REGION Network 2
   RUNG wire#powerrail
      { S7_GenerateENO := "TRUE" } Move(in := "1#煤粉仓2#温度":P, out1 => "MNL"."1#煤粉仓2#温度")
   END_RUNG
   // the same network as SCL:
   "MNL"."1#煤粉仓2#温度" := "1#煤粉仓2#温度":P;
END_REGION

REGION Network 3
   RUNG wire#powerrail
      { S7_GenerateENO := "TRUE" } Move(in := "1#煤粉仓3#温度":P, out1 => "MNL"."1#煤粉仓3#温度")
   END_RUNG
   // the same network as SCL:
   "MNL"."1#煤粉仓3#温度" := "1#煤粉仓3#温度":P;
END_REGION

REGION Network 4
   RUNG wire#powerrail
      { S7_GenerateENO := "TRUE" } Move(in := "Tag_101":P, out1 => "MNL"."1#煤粉仓4#温度")
   END_RUNG
   // the same network as SCL:
   "MNL"."1#煤粉仓4#温度" := "Tag_101":P;
END_REGION

REGION Network 5
   RUNG wire#powerrail
      { S7_GenerateENO := "TRUE" } Move(in := "1#煤粉仓5#温度":P, out1 => "MNL"."1#煤粉仓5#温度")
   END_RUNG
   // the same network as SCL:
   "MNL"."1#煤粉仓5#温度" := "1#煤粉仓5#温度":P;
END_REGION

REGION Network 6
   RUNG wire#powerrail
      { S7_GenerateENO := "TRUE" } Move(in := "1#煤粉仓6#温度":P, out1 => "MNL"."1#煤粉仓6#温度")
   END_RUNG
   // the same network as SCL:
   "MNL"."1#煤粉仓6#温度" := "1#煤粉仓6#温度":P;
END_REGION

REGION Network 7
   RUNG wire#powerrail
      { S7_GenerateENO := "TRUE" } Move(in := "2#煤粉仓1#温度":P, out1 => "MNL"."2#煤粉仓1#温度")
   END_RUNG
   // the same network as SCL:
   "MNL"."2#煤粉仓1#温度" := "2#煤粉仓1#温度":P;
END_REGION

REGION Network 8
   RUNG wire#powerrail
      { S7_GenerateENO := "TRUE" } Move(in := "2#煤粉仓2#温度":P, out1 => "MNL"."2#煤粉仓2#温度")
   END_RUNG
   // the same network as SCL:
   "MNL"."2#煤粉仓2#温度" := "2#煤粉仓2#温度":P;
END_REGION

REGION Network 9
   RUNG wire#powerrail
      { S7_GenerateENO := "TRUE" } Move(in := "2#煤粉仓3#温度":P, out1 => "MNL"."2#煤粉仓3#温度")
   END_RUNG
   // the same network as SCL:
   "MNL"."2#煤粉仓3#温度" := "2#煤粉仓3#温度":P;
END_REGION

REGION Network 10
   RUNG wire#powerrail
      { S7_GenerateENO := "TRUE" } Move(in := "2#煤粉仓4#温度":P, out1 => "MNL"."2#煤粉仓4#温度")
   END_RUNG
   // the same network as SCL:
   "MNL"."2#煤粉仓4#温度" := "2#煤粉仓4#温度":P;
END_REGION

REGION Network 11
   RUNG wire#powerrail
      { S7_GenerateENO := "TRUE" } Move(in := "2#煤粉仓5#温度":P, out1 => "MNL"."2#煤粉仓5#温度")
   END_RUNG
   // the same network as SCL:
   "MNL"."2#煤粉仓5#温度" := "2#煤粉仓5#温度":P;
END_REGION

REGION Network 12
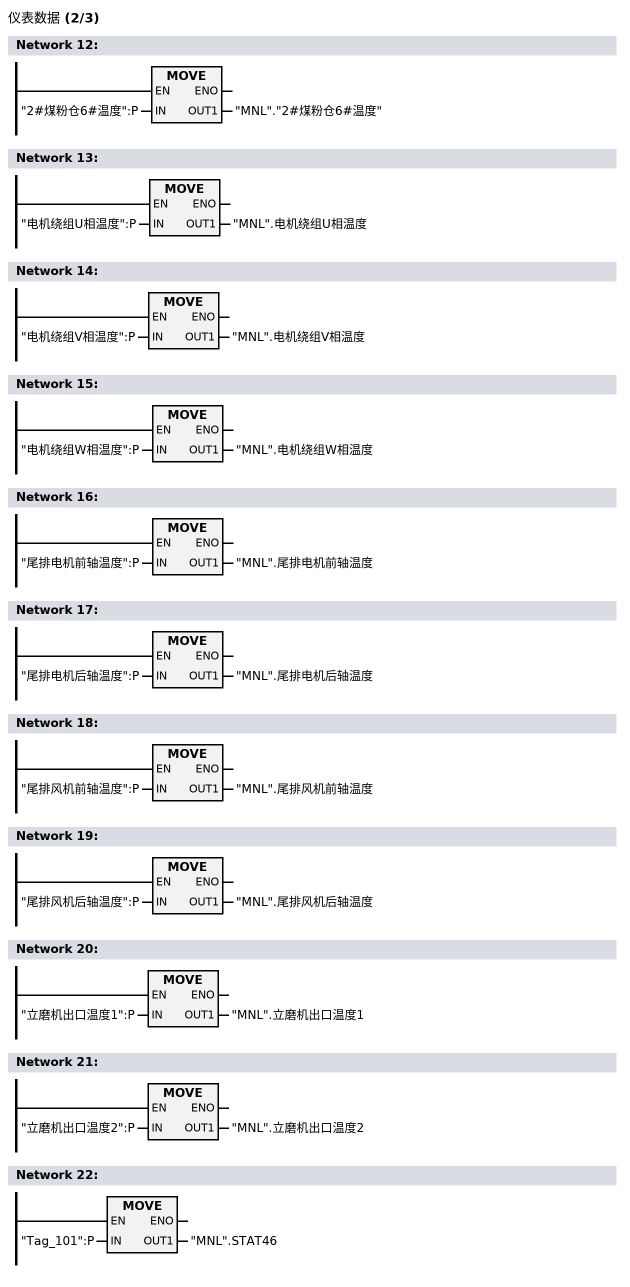
   RUNG wire#powerrail
      { S7_GenerateENO := "TRUE" } Move(in := "2#煤粉仓6#温度":P, out1 => "MNL"."2#煤粉仓6#温度")
   END_RUNG
   // the same network as SCL:
   "MNL"."2#煤粉仓6#温度" := "2#煤粉仓6#温度":P;
END_REGION

REGION Network 13
   RUNG wire#powerrail
      { S7_GenerateENO := "TRUE" } Move(in := "电机绕组U相温度":P, out1 => "MNL".电机绕组U相温度)
   END_RUNG
   // the same network as SCL:
   "MNL".电机绕组U相温度 := "电机绕组U相温度":P;
END_REGION

REGION Network 14
   RUNG wire#powerrail
      { S7_GenerateENO := "TRUE" } Move(in := "电机绕组V相温度":P, out1 => "MNL".电机绕组V相温度)
   END_RUNG
   // the same network as SCL:
   "MNL".电机绕组V相温度 := "电机绕组V相温度":P;
END_REGION

REGION Network 15
   RUNG wire#powerrail
      { S7_GenerateENO := "TRUE" } Move(in := "电机绕组W相温度":P, out1 => "MNL".电机绕组W相温度)
   END_RUNG
   // the same network as SCL:
   "MNL".电机绕组W相温度 := "电机绕组W相温度":P;
END_REGION

REGION Network 16
   RUNG wire#powerrail
      { S7_GenerateENO := "TRUE" } Move(in := "尾排电机前轴温度":P, out1 => "MNL".尾排电机前轴温度)
   END_RUNG
   // the same network as SCL:
   "MNL".尾排电机前轴温度 := "尾排电机前轴温度":P;
END_REGION

REGION Network 17
   RUNG wire#powerrail
      { S7_GenerateENO := "TRUE" } Move(in := "尾排电机后轴温度":P, out1 => "MNL".尾排电机后轴温度)
   END_RUNG
   // the same network as SCL:
   "MNL".尾排电机后轴温度 := "尾排电机后轴温度":P;
END_REGION

REGION Network 18
   RUNG wire#powerrail
      { S7_GenerateENO := "TRUE" } Move(in := "尾排风机前轴温度":P, out1 => "MNL".尾排风机前轴温度)
   END_RUNG
   // the same network as SCL:
   "MNL".尾排风机前轴温度 := "尾排风机前轴温度":P;
END_REGION

REGION Network 19
   RUNG wire#powerrail
      { S7_GenerateENO := "TRUE" } Move(in := "尾排风机后轴温度":P, out1 => "MNL".尾排风机后轴温度)
   END_RUNG
   // the same network as SCL:
   "MNL".尾排风机后轴温度 := "尾排风机后轴温度":P;
END_REGION

REGION Network 20
   RUNG wire#powerrail
      { S7_GenerateENO := "TRUE" } Move(in := "立磨机出口温度1":P, out1 => "MNL".立磨机出口温度1)
   END_RUNG
   // the same network as SCL:
   "MNL".立磨机出口温度1 := "立磨机出口温度1":P;
END_REGION

REGION Network 21
   RUNG wire#powerrail
      { S7_GenerateENO := "TRUE" } Move(in := "立磨机出口温度2":P, out1 => "MNL".立磨机出口温度2)
   END_RUNG
   // the same network as SCL:
   "MNL".立磨机出口温度2 := "立磨机出口温度2":P;
END_REGION

REGION Network 22
   RUNG wire#powerrail
      { S7_GenerateENO := "TRUE" } Move(in := "Tag_101":P, out1 => "MNL".STAT46)
   END_RUNG
   // the same network as SCL:
   "MNL".STAT46 := "Tag_101":P;
END_REGION

REGION Network 23
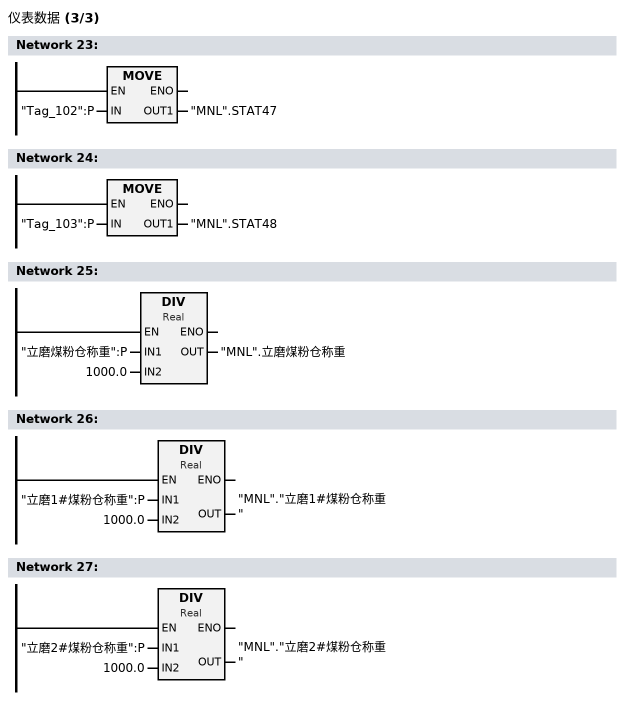
   RUNG wire#powerrail
      { S7_GenerateENO := "TRUE" } Move(in := "Tag_102":P, out1 => "MNL".STAT47)
   END_RUNG
   // the same network as SCL:
   "MNL".STAT47 := "Tag_102":P;
END_REGION

REGION Network 24
   RUNG wire#powerrail
      { S7_GenerateENO := "TRUE" } Move(in := "Tag_103":P, out1 => "MNL".STAT48)
   END_RUNG
   // the same network as SCL:
   "MNL".STAT48 := "Tag_103":P;
END_REGION

REGION Network 25
   RUNG wire#powerrail
      { S7_Templates := "SrcType := Real" } Div(in1 := "立磨煤粉仓称重":P, in2 := 1000.0, out => "MNL".立磨煤粉仓称重)
   END_RUNG
   // the same network as SCL:
   "MNL".立磨煤粉仓称重 := "立磨煤粉仓称重":P / 1000.0;
END_REGION

REGION Network 26
   RUNG wire#powerrail
      { S7_Templates := "SrcType := Real" } Div(in1 := "立磨1#煤粉仓称重":P, in2 := 1000.0, out => "MNL"."立磨1#煤粉仓称重")
   END_RUNG
   // the same network as SCL:
   "MNL"."立磨1#煤粉仓称重" := "立磨1#煤粉仓称重":P / 1000.0;
END_REGION

REGION Network 27
   RUNG wire#powerrail
      { S7_Templates := "SrcType := Real" } Div(in1 := "立磨2#煤粉仓称重":P, in2 := 1000.0, out => "MNL"."立磨2#煤粉仓称重")
   END_RUNG
   // the same network as SCL:
   "MNL"."立磨2#煤粉仓称重" := "立磨2#煤粉仓称重":P / 1000.0;
END_REGION
END_FUNCTION

FUNCTION "NET_RW" : Void   // FC5, LAD
{ S7_Optimized_Access := 'FALSE' }
VERSION : 0.1
BEGIN

REGION Network 1
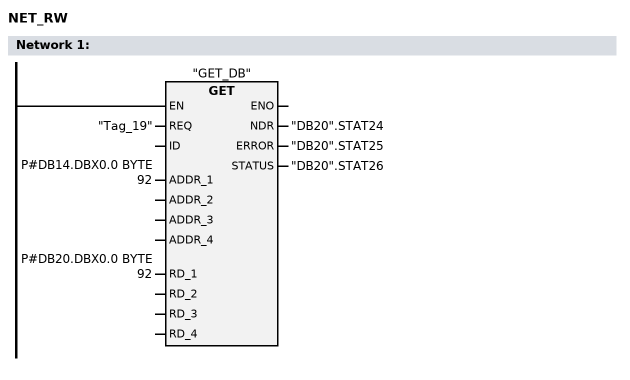
   "GET_DB"(REQ := "Tag_19",   // GET
            ADDR_1 := P#DB14.DBX0.0 BYTE 92,
            RD_1 := P#DB20.DBX0.0 BYTE 92,
            NDR => "DB20".STAT24,
            ERROR => "DB20".STAT25,
            STATUS => "DB20".STAT26);
END_REGION
END_FUNCTION

FUNCTION "仓式泵通信" : Void   // FC6, LAD
{ S7_Optimized_Access := 'TRUE' }
VERSION : 0.1
   VAR_TEMP
      TEMP1 : Bool;
      TEMP2 : Bool;
      TEMP3 : Bool;
      TEMP4 : Bool;
      TEMP5 : Word;
      TEMP6 : Word;
   END_VAR
BEGIN

REGION Network 1
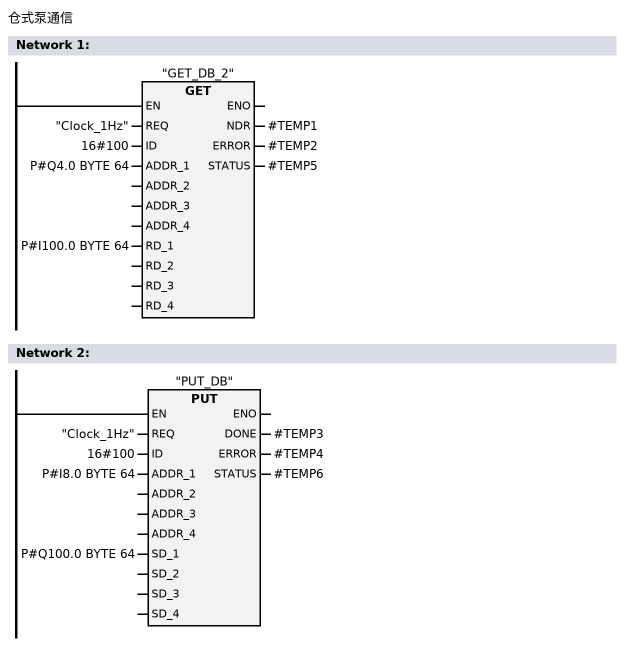
   "GET_DB_2"(REQ := "Clock_1Hz",   // GET
              ID := 16#100,
              ADDR_1 := P#Q4.0 BYTE 64,
              RD_1 := P#I100.0 BYTE 64,
              NDR => #TEMP1,
              ERROR => #TEMP2,
              STATUS => #TEMP5);
END_REGION

REGION Network 2
   "PUT_DB"(REQ := "Clock_1Hz",   // PUT
            ID := 16#100,
            ADDR_1 := P#I8.0 BYTE 64,
            SD_1 := P#Q100.0 BYTE 64,
            DONE => #TEMP3,
            ERROR => #TEMP4,
            STATUS => #TEMP6);
END_REGION
END_FUNCTION

FUNCTION "温度报警输出" : Void   // FC7, LAD
{ S7_Optimized_Access := 'TRUE' }
VERSION : 0.1
   VAR_TEMP   // added for the SCL form of the ladder/FBD networks
      _w1 : Bool;
   END_VAR
BEGIN

REGION Network 1
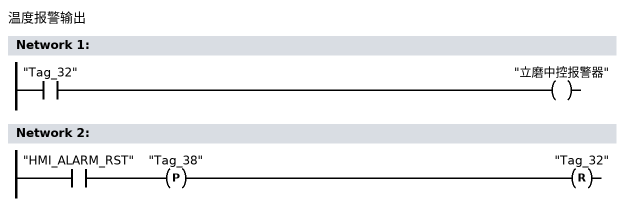
   RUNG wire#powerrail
      Contact( "Tag_32" )
      Coil( "立磨中控报警器" )
   END_RUNG
   // the same network as SCL:
   "立磨中控报警器" := "Tag_32";
END_REGION

REGION Network 2
   RUNG wire#powerrail
      Contact( "HMI_ALARM_RST" )
      P_Trig( "Tag_38" )
      R_Coil( "Tag_32" )
   END_RUNG
   // the same network as SCL:
   #_w1 := "HMI_ALARM_RST" AND NOT "Tag_38";   // rising edge
   "Tag_38" := "HMI_ALARM_RST";
   IF #_w1 THEN "Tag_32" := FALSE; END_IF;
END_REGION
END_FUNCTION

FUNCTION "FC11_DATA_ALARM_FC" : Void   // FC11, LAD
{ S7_Optimized_Access := 'TRUE' }
VERSION : 0.1
   VAR_TEMP   // added for the SCL form of the ladder/FBD networks
      _w1 : Bool;
      _w2 : Bool;
   END_VAR
BEGIN

REGION Network 1
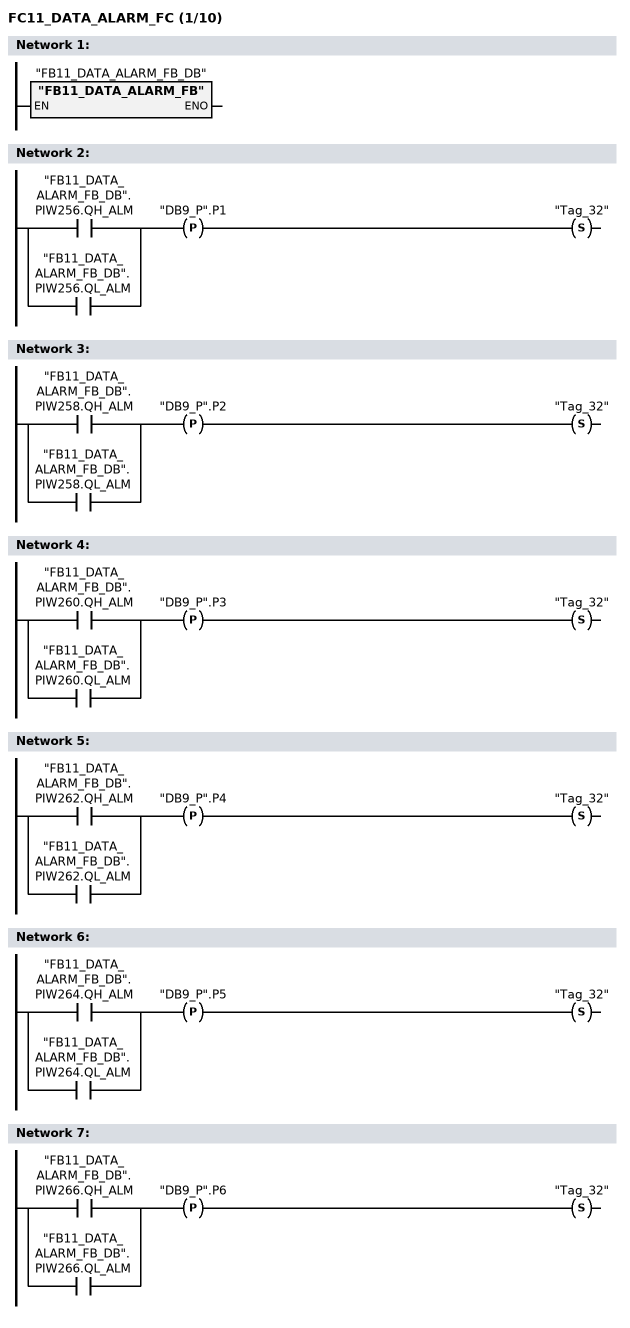
   RUNG wire#powerrail
      "FB11_DATA_ALARM_FB_DB"()
   END_RUNG
   // the same network as SCL:
   "FB11_DATA_ALARM_FB_DB"();   // "FB11_DATA_ALARM_FB"
END_REGION

REGION Network 2
   RUNG wire#powerrail
      Contact( "FB11_DATA_ALARM_FB_DB".PIW256.QH_ALM )
      wire#w1
      P_Trig( "DB9_P".P1 )
      S_Coil( "Tag_32" )
   END_RUNG
   RUNG wire#powerrail
      Contact( "FB11_DATA_ALARM_FB_DB".PIW256.QL_ALM )
   END_RUNG wire#w1
   // the same network as SCL:
   #_w1 := "FB11_DATA_ALARM_FB_DB".PIW256.QH_ALM OR "FB11_DATA_ALARM_FB_DB".PIW256.QL_ALM;
   #_w2 := #_w1 AND NOT "DB9_P".P1;   // rising edge
   "DB9_P".P1 := #_w1;
   IF #_w2 THEN "Tag_32" := TRUE; END_IF;
END_REGION

REGION Network 3
   RUNG wire#powerrail
      Contact( "FB11_DATA_ALARM_FB_DB".PIW258.QH_ALM )
      wire#w1
      P_Trig( "DB9_P".P2 )
      S_Coil( "Tag_32" )
   END_RUNG
   RUNG wire#powerrail
      Contact( "FB11_DATA_ALARM_FB_DB".PIW258.QL_ALM )
   END_RUNG wire#w1
   // the same network as SCL:
   #_w1 := "FB11_DATA_ALARM_FB_DB".PIW258.QH_ALM OR "FB11_DATA_ALARM_FB_DB".PIW258.QL_ALM;
   #_w2 := #_w1 AND NOT "DB9_P".P2;   // rising edge
   "DB9_P".P2 := #_w1;
   IF #_w2 THEN "Tag_32" := TRUE; END_IF;
END_REGION

REGION Network 4
   RUNG wire#powerrail
      Contact( "FB11_DATA_ALARM_FB_DB".PIW260.QH_ALM )
      wire#w1
      P_Trig( "DB9_P".P3 )
      S_Coil( "Tag_32" )
   END_RUNG
   RUNG wire#powerrail
      Contact( "FB11_DATA_ALARM_FB_DB".PIW260.QL_ALM )
   END_RUNG wire#w1
   // the same network as SCL:
   #_w1 := "FB11_DATA_ALARM_FB_DB".PIW260.QH_ALM OR "FB11_DATA_ALARM_FB_DB".PIW260.QL_ALM;
   #_w2 := #_w1 AND NOT "DB9_P".P3;   // rising edge
   "DB9_P".P3 := #_w1;
   IF #_w2 THEN "Tag_32" := TRUE; END_IF;
END_REGION

REGION Network 5
   RUNG wire#powerrail
      Contact( "FB11_DATA_ALARM_FB_DB".PIW262.QH_ALM )
      wire#w1
      P_Trig( "DB9_P".P4 )
      S_Coil( "Tag_32" )
   END_RUNG
   RUNG wire#powerrail
      Contact( "FB11_DATA_ALARM_FB_DB".PIW262.QL_ALM )
   END_RUNG wire#w1
   // the same network as SCL:
   #_w1 := "FB11_DATA_ALARM_FB_DB".PIW262.QH_ALM OR "FB11_DATA_ALARM_FB_DB".PIW262.QL_ALM;
   #_w2 := #_w1 AND NOT "DB9_P".P4;   // rising edge
   "DB9_P".P4 := #_w1;
   IF #_w2 THEN "Tag_32" := TRUE; END_IF;
END_REGION

REGION Network 6
   RUNG wire#powerrail
      Contact( "FB11_DATA_ALARM_FB_DB".PIW264.QH_ALM )
      wire#w1
      P_Trig( "DB9_P".P5 )
      S_Coil( "Tag_32" )
   END_RUNG
   RUNG wire#powerrail
      Contact( "FB11_DATA_ALARM_FB_DB".PIW264.QL_ALM )
   END_RUNG wire#w1
   // the same network as SCL:
   #_w1 := "FB11_DATA_ALARM_FB_DB".PIW264.QH_ALM OR "FB11_DATA_ALARM_FB_DB".PIW264.QL_ALM;
   #_w2 := #_w1 AND NOT "DB9_P".P5;   // rising edge
   "DB9_P".P5 := #_w1;
   IF #_w2 THEN "Tag_32" := TRUE; END_IF;
END_REGION

REGION Network 7
   RUNG wire#powerrail
      Contact( "FB11_DATA_ALARM_FB_DB".PIW266.QH_ALM )
      wire#w1
      P_Trig( "DB9_P".P6 )
      S_Coil( "Tag_32" )
   END_RUNG
   RUNG wire#powerrail
      Contact( "FB11_DATA_ALARM_FB_DB".PIW266.QL_ALM )
   END_RUNG wire#w1
   // the same network as SCL:
   #_w1 := "FB11_DATA_ALARM_FB_DB".PIW266.QH_ALM OR "FB11_DATA_ALARM_FB_DB".PIW266.QL_ALM;
   #_w2 := #_w1 AND NOT "DB9_P".P6;   // rising edge
   "DB9_P".P6 := #_w1;
   IF #_w2 THEN "Tag_32" := TRUE; END_IF;
END_REGION

REGION Network 8
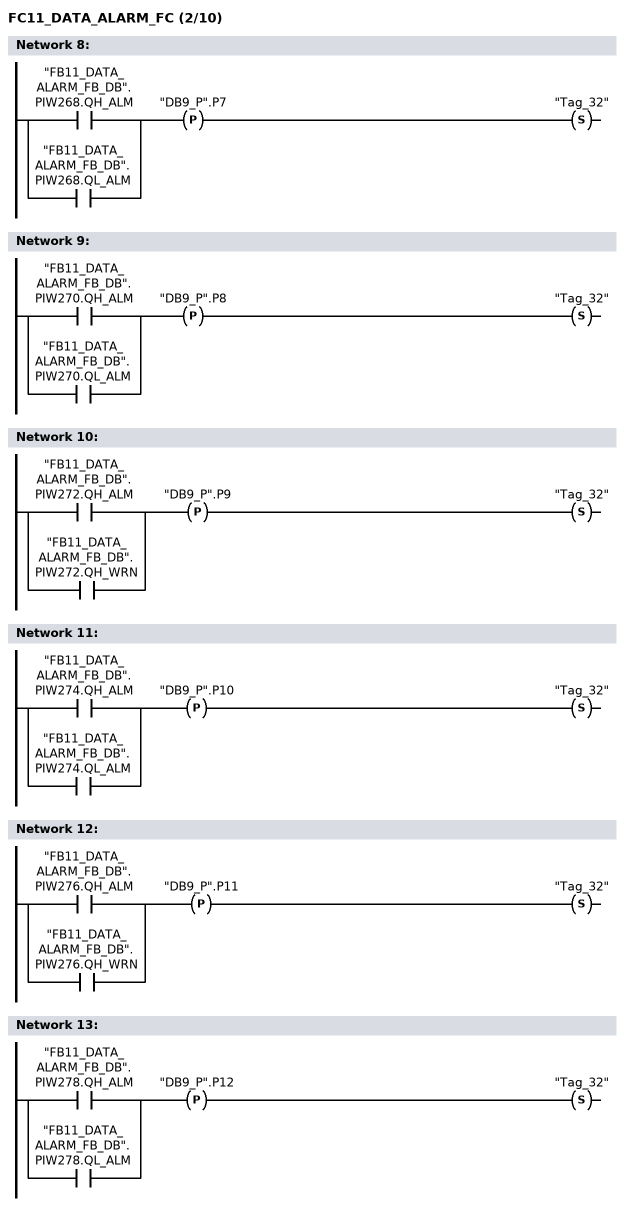
   RUNG wire#powerrail
      Contact( "FB11_DATA_ALARM_FB_DB".PIW268.QH_ALM )
      wire#w1
      P_Trig( "DB9_P".P7 )
      S_Coil( "Tag_32" )
   END_RUNG
   RUNG wire#powerrail
      Contact( "FB11_DATA_ALARM_FB_DB".PIW268.QL_ALM )
   END_RUNG wire#w1
   // the same network as SCL:
   #_w1 := "FB11_DATA_ALARM_FB_DB".PIW268.QH_ALM OR "FB11_DATA_ALARM_FB_DB".PIW268.QL_ALM;
   #_w2 := #_w1 AND NOT "DB9_P".P7;   // rising edge
   "DB9_P".P7 := #_w1;
   IF #_w2 THEN "Tag_32" := TRUE; END_IF;
END_REGION

REGION Network 9
   RUNG wire#powerrail
      Contact( "FB11_DATA_ALARM_FB_DB".PIW270.QH_ALM )
      wire#w1
      P_Trig( "DB9_P".P8 )
      S_Coil( "Tag_32" )
   END_RUNG
   RUNG wire#powerrail
      Contact( "FB11_DATA_ALARM_FB_DB".PIW270.QL_ALM )
   END_RUNG wire#w1
   // the same network as SCL:
   #_w1 := "FB11_DATA_ALARM_FB_DB".PIW270.QH_ALM OR "FB11_DATA_ALARM_FB_DB".PIW270.QL_ALM;
   #_w2 := #_w1 AND NOT "DB9_P".P8;   // rising edge
   "DB9_P".P8 := #_w1;
   IF #_w2 THEN "Tag_32" := TRUE; END_IF;
END_REGION

REGION Network 10
   RUNG wire#powerrail
      Contact( "FB11_DATA_ALARM_FB_DB".PIW272.QH_ALM )
      wire#w1
      P_Trig( "DB9_P".P9 )
      S_Coil( "Tag_32" )
   END_RUNG
   RUNG wire#powerrail
      Contact( "FB11_DATA_ALARM_FB_DB".PIW272.QH_WRN )
   END_RUNG wire#w1
   // the same network as SCL:
   #_w1 := "FB11_DATA_ALARM_FB_DB".PIW272.QH_ALM OR "FB11_DATA_ALARM_FB_DB".PIW272.QH_WRN;
   #_w2 := #_w1 AND NOT "DB9_P".P9;   // rising edge
   "DB9_P".P9 := #_w1;
   IF #_w2 THEN "Tag_32" := TRUE; END_IF;
END_REGION

REGION Network 11
   RUNG wire#powerrail
      Contact( "FB11_DATA_ALARM_FB_DB".PIW274.QH_ALM )
      wire#w1
      P_Trig( "DB9_P".P10 )
      S_Coil( "Tag_32" )
   END_RUNG
   RUNG wire#powerrail
      Contact( "FB11_DATA_ALARM_FB_DB".PIW274.QL_ALM )
   END_RUNG wire#w1
   // the same network as SCL:
   #_w1 := "FB11_DATA_ALARM_FB_DB".PIW274.QH_ALM OR "FB11_DATA_ALARM_FB_DB".PIW274.QL_ALM;
   #_w2 := #_w1 AND NOT "DB9_P".P10;   // rising edge
   "DB9_P".P10 := #_w1;
   IF #_w2 THEN "Tag_32" := TRUE; END_IF;
END_REGION

REGION Network 12
   RUNG wire#powerrail
      Contact( "FB11_DATA_ALARM_FB_DB".PIW276.QH_ALM )
      wire#w1
      P_Trig( "DB9_P".P11 )
      S_Coil( "Tag_32" )
   END_RUNG
   RUNG wire#powerrail
      Contact( "FB11_DATA_ALARM_FB_DB".PIW276.QH_WRN )
   END_RUNG wire#w1
   // the same network as SCL:
   #_w1 := "FB11_DATA_ALARM_FB_DB".PIW276.QH_ALM OR "FB11_DATA_ALARM_FB_DB".PIW276.QH_WRN;
   #_w2 := #_w1 AND NOT "DB9_P".P11;   // rising edge
   "DB9_P".P11 := #_w1;
   IF #_w2 THEN "Tag_32" := TRUE; END_IF;
END_REGION

REGION Network 13
   RUNG wire#powerrail
      Contact( "FB11_DATA_ALARM_FB_DB".PIW278.QH_ALM )
      wire#w1
      P_Trig( "DB9_P".P12 )
      S_Coil( "Tag_32" )
   END_RUNG
   RUNG wire#powerrail
      Contact( "FB11_DATA_ALARM_FB_DB".PIW278.QL_ALM )
   END_RUNG wire#w1
   // the same network as SCL:
   #_w1 := "FB11_DATA_ALARM_FB_DB".PIW278.QH_ALM OR "FB11_DATA_ALARM_FB_DB".PIW278.QL_ALM;
   #_w2 := #_w1 AND NOT "DB9_P".P12;   // rising edge
   "DB9_P".P12 := #_w1;
   IF #_w2 THEN "Tag_32" := TRUE; END_IF;
END_REGION

REGION Network 14
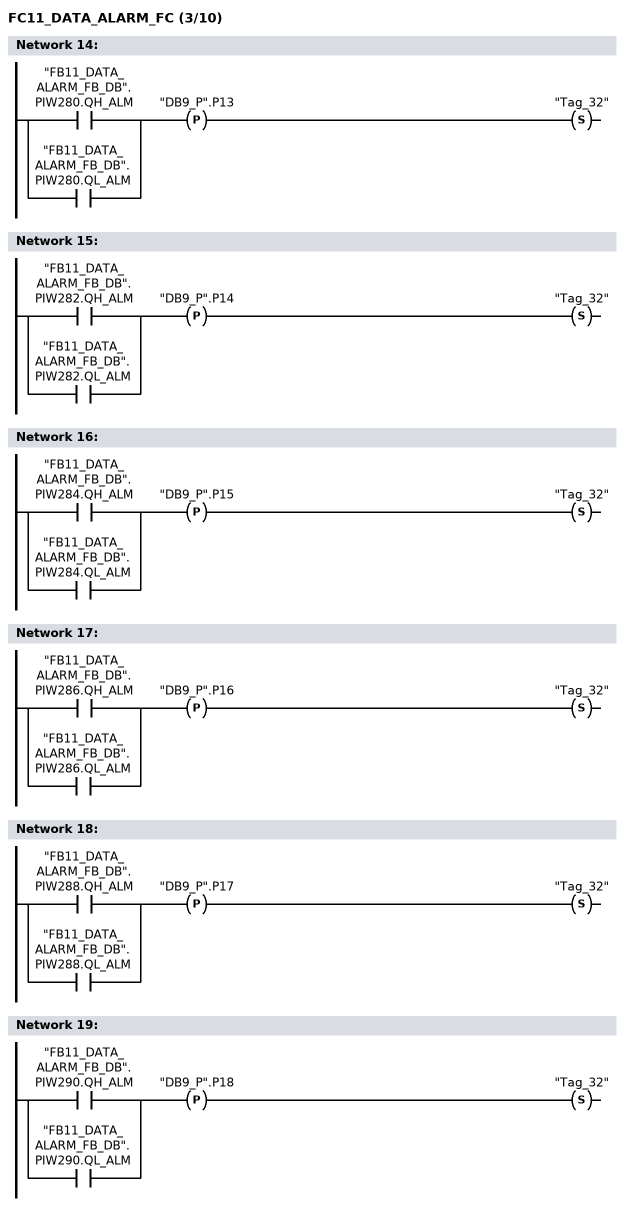
   RUNG wire#powerrail
      Contact( "FB11_DATA_ALARM_FB_DB".PIW280.QH_ALM )
      wire#w1
      P_Trig( "DB9_P".P13 )
      S_Coil( "Tag_32" )
   END_RUNG
   RUNG wire#powerrail
      Contact( "FB11_DATA_ALARM_FB_DB".PIW280.QL_ALM )
   END_RUNG wire#w1
   // the same network as SCL:
   #_w1 := "FB11_DATA_ALARM_FB_DB".PIW280.QH_ALM OR "FB11_DATA_ALARM_FB_DB".PIW280.QL_ALM;
   #_w2 := #_w1 AND NOT "DB9_P".P13;   // rising edge
   "DB9_P".P13 := #_w1;
   IF #_w2 THEN "Tag_32" := TRUE; END_IF;
END_REGION

REGION Network 15
   RUNG wire#powerrail
      Contact( "FB11_DATA_ALARM_FB_DB".PIW282.QH_ALM )
      wire#w1
      P_Trig( "DB9_P".P14 )
      S_Coil( "Tag_32" )
   END_RUNG
   RUNG wire#powerrail
      Contact( "FB11_DATA_ALARM_FB_DB".PIW282.QL_ALM )
   END_RUNG wire#w1
   // the same network as SCL:
   #_w1 := "FB11_DATA_ALARM_FB_DB".PIW282.QH_ALM OR "FB11_DATA_ALARM_FB_DB".PIW282.QL_ALM;
   #_w2 := #_w1 AND NOT "DB9_P".P14;   // rising edge
   "DB9_P".P14 := #_w1;
   IF #_w2 THEN "Tag_32" := TRUE; END_IF;
END_REGION

REGION Network 16
   RUNG wire#powerrail
      Contact( "FB11_DATA_ALARM_FB_DB".PIW284.QH_ALM )
      wire#w1
      P_Trig( "DB9_P".P15 )
      S_Coil( "Tag_32" )
   END_RUNG
   RUNG wire#powerrail
      Contact( "FB11_DATA_ALARM_FB_DB".PIW284.QL_ALM )
   END_RUNG wire#w1
   // the same network as SCL:
   #_w1 := "FB11_DATA_ALARM_FB_DB".PIW284.QH_ALM OR "FB11_DATA_ALARM_FB_DB".PIW284.QL_ALM;
   #_w2 := #_w1 AND NOT "DB9_P".P15;   // rising edge
   "DB9_P".P15 := #_w1;
   IF #_w2 THEN "Tag_32" := TRUE; END_IF;
END_REGION

REGION Network 17
   RUNG wire#powerrail
      Contact( "FB11_DATA_ALARM_FB_DB".PIW286.QH_ALM )
      wire#w1
      P_Trig( "DB9_P".P16 )
      S_Coil( "Tag_32" )
   END_RUNG
   RUNG wire#powerrail
      Contact( "FB11_DATA_ALARM_FB_DB".PIW286.QL_ALM )
   END_RUNG wire#w1
   // the same network as SCL:
   #_w1 := "FB11_DATA_ALARM_FB_DB".PIW286.QH_ALM OR "FB11_DATA_ALARM_FB_DB".PIW286.QL_ALM;
   #_w2 := #_w1 AND NOT "DB9_P".P16;   // rising edge
   "DB9_P".P16 := #_w1;
   IF #_w2 THEN "Tag_32" := TRUE; END_IF;
END_REGION

REGION Network 18
   RUNG wire#powerrail
      Contact( "FB11_DATA_ALARM_FB_DB".PIW288.QH_ALM )
      wire#w1
      P_Trig( "DB9_P".P17 )
      S_Coil( "Tag_32" )
   END_RUNG
   RUNG wire#powerrail
      Contact( "FB11_DATA_ALARM_FB_DB".PIW288.QL_ALM )
   END_RUNG wire#w1
   // the same network as SCL:
   #_w1 := "FB11_DATA_ALARM_FB_DB".PIW288.QH_ALM OR "FB11_DATA_ALARM_FB_DB".PIW288.QL_ALM;
   #_w2 := #_w1 AND NOT "DB9_P".P17;   // rising edge
   "DB9_P".P17 := #_w1;
   IF #_w2 THEN "Tag_32" := TRUE; END_IF;
END_REGION

REGION Network 19
   RUNG wire#powerrail
      Contact( "FB11_DATA_ALARM_FB_DB".PIW290.QH_ALM )
      wire#w1
      P_Trig( "DB9_P".P18 )
      S_Coil( "Tag_32" )
   END_RUNG
   RUNG wire#powerrail
      Contact( "FB11_DATA_ALARM_FB_DB".PIW290.QL_ALM )
   END_RUNG wire#w1
   // the same network as SCL:
   #_w1 := "FB11_DATA_ALARM_FB_DB".PIW290.QH_ALM OR "FB11_DATA_ALARM_FB_DB".PIW290.QL_ALM;
   #_w2 := #_w1 AND NOT "DB9_P".P18;   // rising edge
   "DB9_P".P18 := #_w1;
   IF #_w2 THEN "Tag_32" := TRUE; END_IF;
END_REGION

REGION Network 20
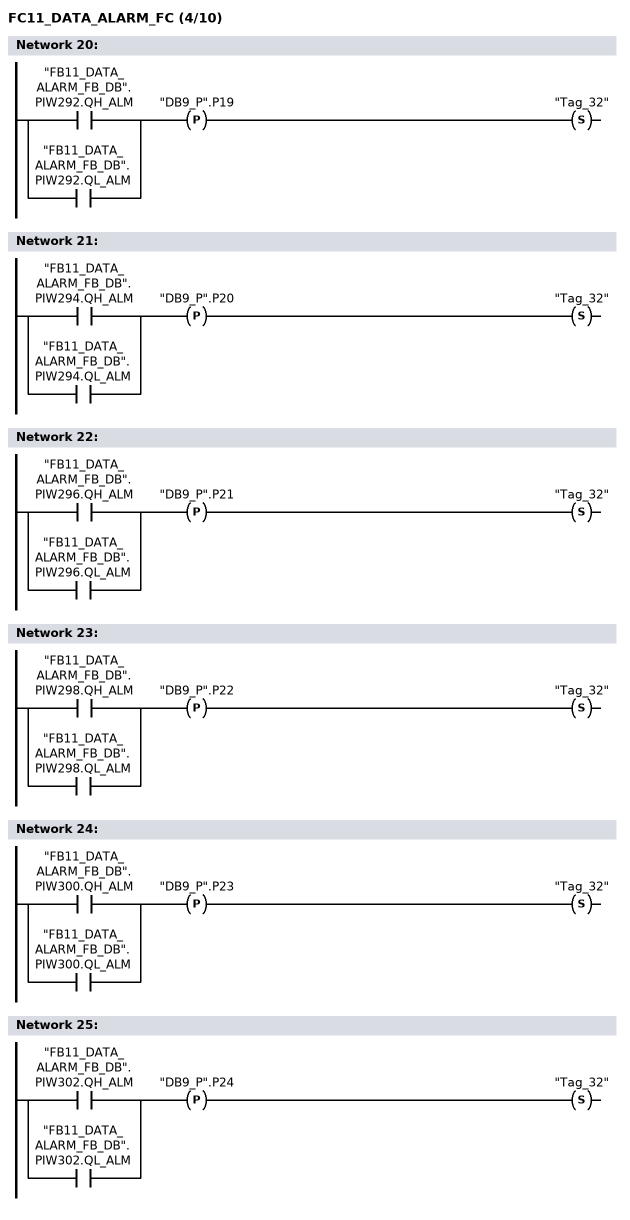
   RUNG wire#powerrail
      Contact( "FB11_DATA_ALARM_FB_DB".PIW292.QH_ALM )
      wire#w1
      P_Trig( "DB9_P".P19 )
      S_Coil( "Tag_32" )
   END_RUNG
   RUNG wire#powerrail
      Contact( "FB11_DATA_ALARM_FB_DB".PIW292.QL_ALM )
   END_RUNG wire#w1
   // the same network as SCL:
   #_w1 := "FB11_DATA_ALARM_FB_DB".PIW292.QH_ALM OR "FB11_DATA_ALARM_FB_DB".PIW292.QL_ALM;
   #_w2 := #_w1 AND NOT "DB9_P".P19;   // rising edge
   "DB9_P".P19 := #_w1;
   IF #_w2 THEN "Tag_32" := TRUE; END_IF;
END_REGION

REGION Network 21
   RUNG wire#powerrail
      Contact( "FB11_DATA_ALARM_FB_DB".PIW294.QH_ALM )
      wire#w1
      P_Trig( "DB9_P".P20 )
      S_Coil( "Tag_32" )
   END_RUNG
   RUNG wire#powerrail
      Contact( "FB11_DATA_ALARM_FB_DB".PIW294.QL_ALM )
   END_RUNG wire#w1
   // the same network as SCL:
   #_w1 := "FB11_DATA_ALARM_FB_DB".PIW294.QH_ALM OR "FB11_DATA_ALARM_FB_DB".PIW294.QL_ALM;
   #_w2 := #_w1 AND NOT "DB9_P".P20;   // rising edge
   "DB9_P".P20 := #_w1;
   IF #_w2 THEN "Tag_32" := TRUE; END_IF;
END_REGION

REGION Network 22
   RUNG wire#powerrail
      Contact( "FB11_DATA_ALARM_FB_DB".PIW296.QH_ALM )
      wire#w1
      P_Trig( "DB9_P".P21 )
      S_Coil( "Tag_32" )
   END_RUNG
   RUNG wire#powerrail
      Contact( "FB11_DATA_ALARM_FB_DB".PIW296.QL_ALM )
   END_RUNG wire#w1
   // the same network as SCL:
   #_w1 := "FB11_DATA_ALARM_FB_DB".PIW296.QH_ALM OR "FB11_DATA_ALARM_FB_DB".PIW296.QL_ALM;
   #_w2 := #_w1 AND NOT "DB9_P".P21;   // rising edge
   "DB9_P".P21 := #_w1;
   IF #_w2 THEN "Tag_32" := TRUE; END_IF;
END_REGION

REGION Network 23
   RUNG wire#powerrail
      Contact( "FB11_DATA_ALARM_FB_DB".PIW298.QH_ALM )
      wire#w1
      P_Trig( "DB9_P".P22 )
      S_Coil( "Tag_32" )
   END_RUNG
   RUNG wire#powerrail
      Contact( "FB11_DATA_ALARM_FB_DB".PIW298.QL_ALM )
   END_RUNG wire#w1
   // the same network as SCL:
   #_w1 := "FB11_DATA_ALARM_FB_DB".PIW298.QH_ALM OR "FB11_DATA_ALARM_FB_DB".PIW298.QL_ALM;
   #_w2 := #_w1 AND NOT "DB9_P".P22;   // rising edge
   "DB9_P".P22 := #_w1;
   IF #_w2 THEN "Tag_32" := TRUE; END_IF;
END_REGION

REGION Network 24
   RUNG wire#powerrail
      Contact( "FB11_DATA_ALARM_FB_DB".PIW300.QH_ALM )
      wire#w1
      P_Trig( "DB9_P".P23 )
      S_Coil( "Tag_32" )
   END_RUNG
   RUNG wire#powerrail
      Contact( "FB11_DATA_ALARM_FB_DB".PIW300.QL_ALM )
   END_RUNG wire#w1
   // the same network as SCL:
   #_w1 := "FB11_DATA_ALARM_FB_DB".PIW300.QH_ALM OR "FB11_DATA_ALARM_FB_DB".PIW300.QL_ALM;
   #_w2 := #_w1 AND NOT "DB9_P".P23;   // rising edge
   "DB9_P".P23 := #_w1;
   IF #_w2 THEN "Tag_32" := TRUE; END_IF;
END_REGION

REGION Network 25
   RUNG wire#powerrail
      Contact( "FB11_DATA_ALARM_FB_DB".PIW302.QH_ALM )
      wire#w1
      P_Trig( "DB9_P".P24 )
      S_Coil( "Tag_32" )
   END_RUNG
   RUNG wire#powerrail
      Contact( "FB11_DATA_ALARM_FB_DB".PIW302.QL_ALM )
   END_RUNG wire#w1
   // the same network as SCL:
   #_w1 := "FB11_DATA_ALARM_FB_DB".PIW302.QH_ALM OR "FB11_DATA_ALARM_FB_DB".PIW302.QL_ALM;
   #_w2 := #_w1 AND NOT "DB9_P".P24;   // rising edge
   "DB9_P".P24 := #_w1;
   IF #_w2 THEN "Tag_32" := TRUE; END_IF;
END_REGION

REGION Network 26
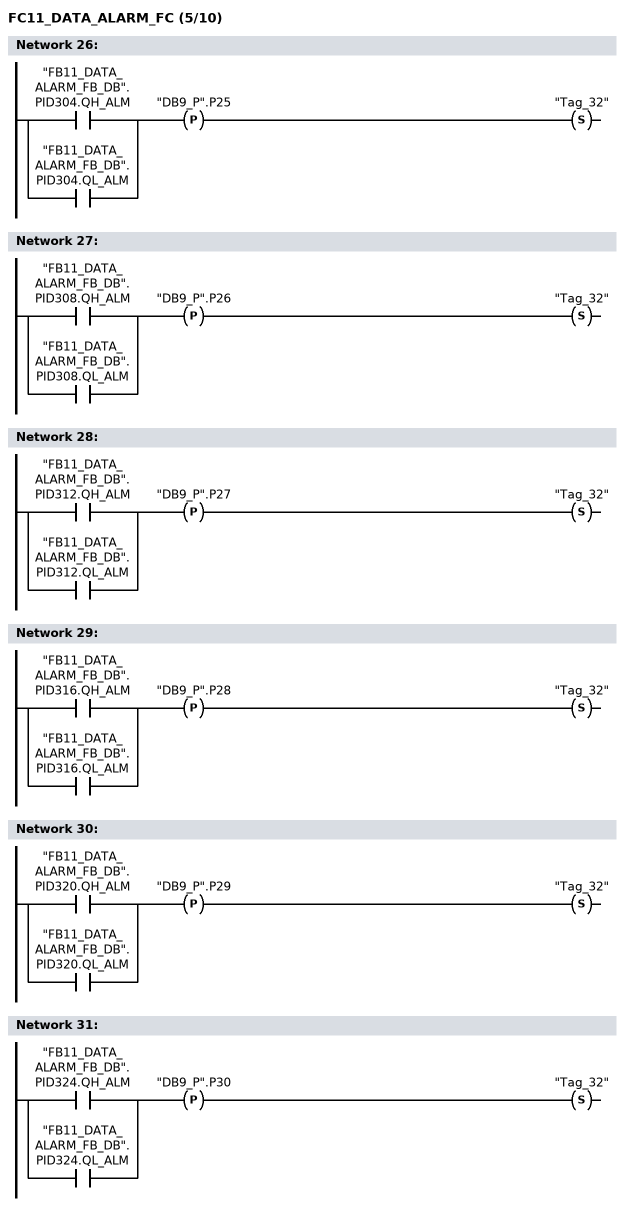
   RUNG wire#powerrail
      Contact( "FB11_DATA_ALARM_FB_DB".PID304.QH_ALM )
      wire#w1
      P_Trig( "DB9_P".P25 )
      S_Coil( "Tag_32" )
   END_RUNG
   RUNG wire#powerrail
      Contact( "FB11_DATA_ALARM_FB_DB".PID304.QL_ALM )
   END_RUNG wire#w1
   // the same network as SCL:
   #_w1 := "FB11_DATA_ALARM_FB_DB".PID304.QH_ALM OR "FB11_DATA_ALARM_FB_DB".PID304.QL_ALM;
   #_w2 := #_w1 AND NOT "DB9_P".P25;   // rising edge
   "DB9_P".P25 := #_w1;
   IF #_w2 THEN "Tag_32" := TRUE; END_IF;
END_REGION

REGION Network 27
   RUNG wire#powerrail
      Contact( "FB11_DATA_ALARM_FB_DB".PID308.QH_ALM )
      wire#w1
      P_Trig( "DB9_P".P26 )
      S_Coil( "Tag_32" )
   END_RUNG
   RUNG wire#powerrail
      Contact( "FB11_DATA_ALARM_FB_DB".PID308.QL_ALM )
   END_RUNG wire#w1
   // the same network as SCL:
   #_w1 := "FB11_DATA_ALARM_FB_DB".PID308.QH_ALM OR "FB11_DATA_ALARM_FB_DB".PID308.QL_ALM;
   #_w2 := #_w1 AND NOT "DB9_P".P26;   // rising edge
   "DB9_P".P26 := #_w1;
   IF #_w2 THEN "Tag_32" := TRUE; END_IF;
END_REGION

REGION Network 28
   RUNG wire#powerrail
      Contact( "FB11_DATA_ALARM_FB_DB".PID312.QH_ALM )
      wire#w1
      P_Trig( "DB9_P".P27 )
      S_Coil( "Tag_32" )
   END_RUNG
   RUNG wire#powerrail
      Contact( "FB11_DATA_ALARM_FB_DB".PID312.QL_ALM )
   END_RUNG wire#w1
   // the same network as SCL:
   #_w1 := "FB11_DATA_ALARM_FB_DB".PID312.QH_ALM OR "FB11_DATA_ALARM_FB_DB".PID312.QL_ALM;
   #_w2 := #_w1 AND NOT "DB9_P".P27;   // rising edge
   "DB9_P".P27 := #_w1;
   IF #_w2 THEN "Tag_32" := TRUE; END_IF;
END_REGION

REGION Network 29
   RUNG wire#powerrail
      Contact( "FB11_DATA_ALARM_FB_DB".PID316.QH_ALM )
      wire#w1
      P_Trig( "DB9_P".P28 )
      S_Coil( "Tag_32" )
   END_RUNG
   RUNG wire#powerrail
      Contact( "FB11_DATA_ALARM_FB_DB".PID316.QL_ALM )
   END_RUNG wire#w1
   // the same network as SCL:
   #_w1 := "FB11_DATA_ALARM_FB_DB".PID316.QH_ALM OR "FB11_DATA_ALARM_FB_DB".PID316.QL_ALM;
   #_w2 := #_w1 AND NOT "DB9_P".P28;   // rising edge
   "DB9_P".P28 := #_w1;
   IF #_w2 THEN "Tag_32" := TRUE; END_IF;
END_REGION

REGION Network 30
   RUNG wire#powerrail
      Contact( "FB11_DATA_ALARM_FB_DB".PID320.QH_ALM )
      wire#w1
      P_Trig( "DB9_P".P29 )
      S_Coil( "Tag_32" )
   END_RUNG
   RUNG wire#powerrail
      Contact( "FB11_DATA_ALARM_FB_DB".PID320.QL_ALM )
   END_RUNG wire#w1
   // the same network as SCL:
   #_w1 := "FB11_DATA_ALARM_FB_DB".PID320.QH_ALM OR "FB11_DATA_ALARM_FB_DB".PID320.QL_ALM;
   #_w2 := #_w1 AND NOT "DB9_P".P29;   // rising edge
   "DB9_P".P29 := #_w1;
   IF #_w2 THEN "Tag_32" := TRUE; END_IF;
END_REGION

REGION Network 31
   RUNG wire#powerrail
      Contact( "FB11_DATA_ALARM_FB_DB".PID324.QH_ALM )
      wire#w1
      P_Trig( "DB9_P".P30 )
      S_Coil( "Tag_32" )
   END_RUNG
   RUNG wire#powerrail
      Contact( "FB11_DATA_ALARM_FB_DB".PID324.QL_ALM )
   END_RUNG wire#w1
   // the same network as SCL:
   #_w1 := "FB11_DATA_ALARM_FB_DB".PID324.QH_ALM OR "FB11_DATA_ALARM_FB_DB".PID324.QL_ALM;
   #_w2 := #_w1 AND NOT "DB9_P".P30;   // rising edge
   "DB9_P".P30 := #_w1;
   IF #_w2 THEN "Tag_32" := TRUE; END_IF;
END_REGION

REGION Network 32
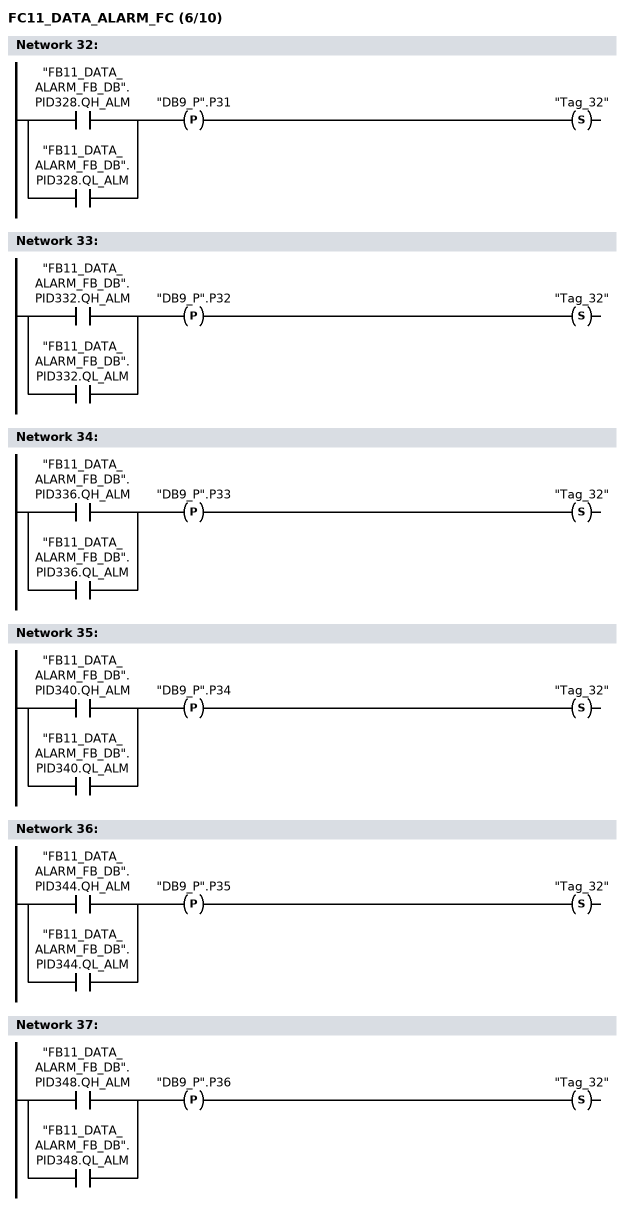
   RUNG wire#powerrail
      Contact( "FB11_DATA_ALARM_FB_DB".PID328.QH_ALM )
      wire#w1
      P_Trig( "DB9_P".P31 )
      S_Coil( "Tag_32" )
   END_RUNG
   RUNG wire#powerrail
      Contact( "FB11_DATA_ALARM_FB_DB".PID328.QL_ALM )
   END_RUNG wire#w1
   // the same network as SCL:
   #_w1 := "FB11_DATA_ALARM_FB_DB".PID328.QH_ALM OR "FB11_DATA_ALARM_FB_DB".PID328.QL_ALM;
   #_w2 := #_w1 AND NOT "DB9_P".P31;   // rising edge
   "DB9_P".P31 := #_w1;
   IF #_w2 THEN "Tag_32" := TRUE; END_IF;
END_REGION

REGION Network 33
   RUNG wire#powerrail
      Contact( "FB11_DATA_ALARM_FB_DB".PID332.QH_ALM )
      wire#w1
      P_Trig( "DB9_P".P32 )
      S_Coil( "Tag_32" )
   END_RUNG
   RUNG wire#powerrail
      Contact( "FB11_DATA_ALARM_FB_DB".PID332.QL_ALM )
   END_RUNG wire#w1
   // the same network as SCL:
   #_w1 := "FB11_DATA_ALARM_FB_DB".PID332.QH_ALM OR "FB11_DATA_ALARM_FB_DB".PID332.QL_ALM;
   #_w2 := #_w1 AND NOT "DB9_P".P32;   // rising edge
   "DB9_P".P32 := #_w1;
   IF #_w2 THEN "Tag_32" := TRUE; END_IF;
END_REGION

REGION Network 34
   RUNG wire#powerrail
      Contact( "FB11_DATA_ALARM_FB_DB".PID336.QH_ALM )
      wire#w1
      P_Trig( "DB9_P".P33 )
      S_Coil( "Tag_32" )
   END_RUNG
   RUNG wire#powerrail
      Contact( "FB11_DATA_ALARM_FB_DB".PID336.QL_ALM )
   END_RUNG wire#w1
   // the same network as SCL:
   #_w1 := "FB11_DATA_ALARM_FB_DB".PID336.QH_ALM OR "FB11_DATA_ALARM_FB_DB".PID336.QL_ALM;
   #_w2 := #_w1 AND NOT "DB9_P".P33;   // rising edge
   "DB9_P".P33 := #_w1;
   IF #_w2 THEN "Tag_32" := TRUE; END_IF;
END_REGION

REGION Network 35
   RUNG wire#powerrail
      Contact( "FB11_DATA_ALARM_FB_DB".PID340.QH_ALM )
      wire#w1
      P_Trig( "DB9_P".P34 )
      S_Coil( "Tag_32" )
   END_RUNG
   RUNG wire#powerrail
      Contact( "FB11_DATA_ALARM_FB_DB".PID340.QL_ALM )
   END_RUNG wire#w1
   // the same network as SCL:
   #_w1 := "FB11_DATA_ALARM_FB_DB".PID340.QH_ALM OR "FB11_DATA_ALARM_FB_DB".PID340.QL_ALM;
   #_w2 := #_w1 AND NOT "DB9_P".P34;   // rising edge
   "DB9_P".P34 := #_w1;
   IF #_w2 THEN "Tag_32" := TRUE; END_IF;
END_REGION

REGION Network 36
   RUNG wire#powerrail
      Contact( "FB11_DATA_ALARM_FB_DB".PID344.QH_ALM )
      wire#w1
      P_Trig( "DB9_P".P35 )
      S_Coil( "Tag_32" )
   END_RUNG
   RUNG wire#powerrail
      Contact( "FB11_DATA_ALARM_FB_DB".PID344.QL_ALM )
   END_RUNG wire#w1
   // the same network as SCL:
   #_w1 := "FB11_DATA_ALARM_FB_DB".PID344.QH_ALM OR "FB11_DATA_ALARM_FB_DB".PID344.QL_ALM;
   #_w2 := #_w1 AND NOT "DB9_P".P35;   // rising edge
   "DB9_P".P35 := #_w1;
   IF #_w2 THEN "Tag_32" := TRUE; END_IF;
END_REGION

REGION Network 37
   RUNG wire#powerrail
      Contact( "FB11_DATA_ALARM_FB_DB".PID348.QH_ALM )
      wire#w1
      P_Trig( "DB9_P".P36 )
      S_Coil( "Tag_32" )
   END_RUNG
   RUNG wire#powerrail
      Contact( "FB11_DATA_ALARM_FB_DB".PID348.QL_ALM )
   END_RUNG wire#w1
   // the same network as SCL:
   #_w1 := "FB11_DATA_ALARM_FB_DB".PID348.QH_ALM OR "FB11_DATA_ALARM_FB_DB".PID348.QL_ALM;
   #_w2 := #_w1 AND NOT "DB9_P".P36;   // rising edge
   "DB9_P".P36 := #_w1;
   IF #_w2 THEN "Tag_32" := TRUE; END_IF;
END_REGION

REGION Network 38
